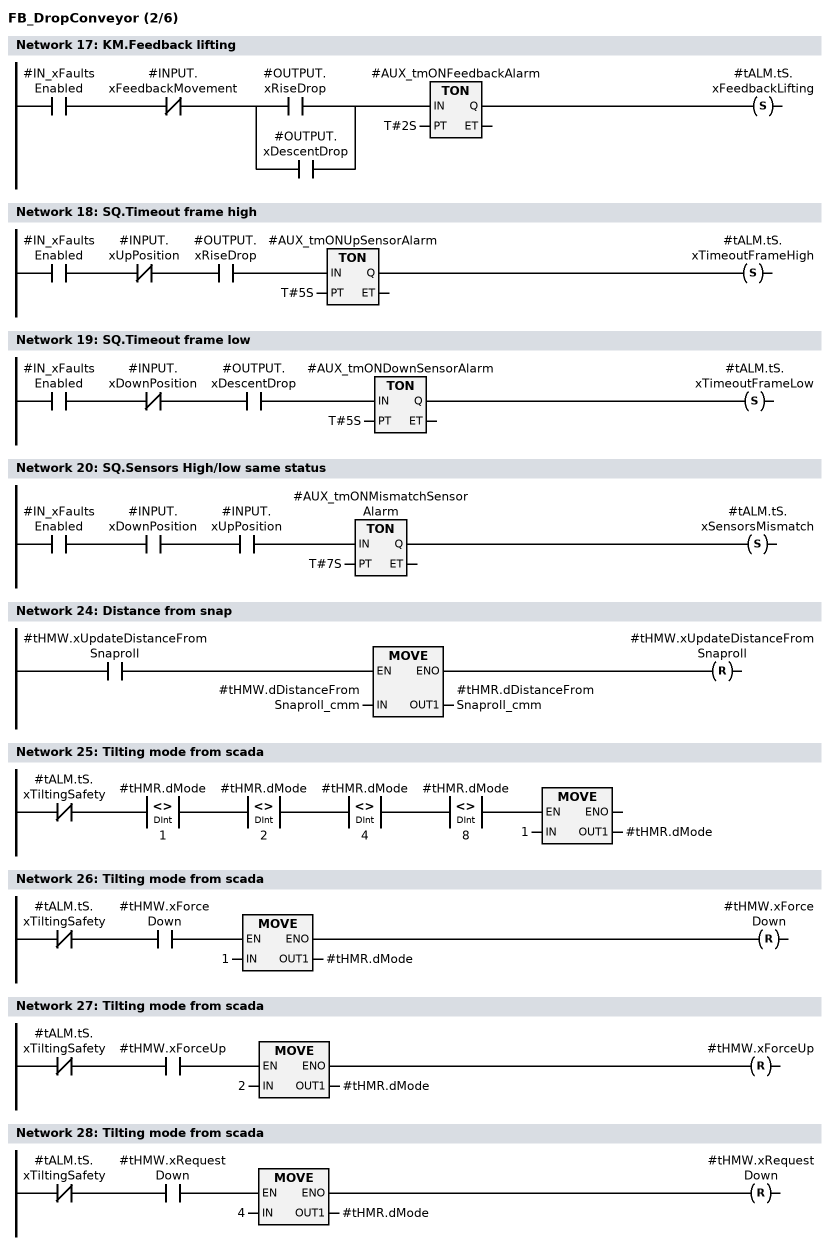
   #AUX_tmONFeedbackAlarm(IN := #IN_xFaultsEnabled AND NOT #INPUT.xFeedbackMovement AND (#OUTPUT.xRiseDrop OR #OUTPUT.xDescentDrop),   // TON
                          PT := T#2S);
   IF #AUX_tmONFeedbackAlarm.Q THEN #tALM.tS.xFeedbackLifting := TRUE; END_IF;
END_REGION

REGION Network 18: SQ.Timeout frame high
   #AUX_tmONUpSensorAlarm(IN := #IN_xFaultsEnabled AND NOT #INPUT.xUpPosition AND #OUTPUT.xRiseDrop, PT := T#5S);   // TON
   IF #AUX_tmONUpSensorAlarm.Q THEN #tALM.tS.xTimeoutFrameHigh := TRUE; END_IF;
END_REGION

REGION Network 19: SQ.Timeout frame low
   #AUX_tmONDownSensorAlarm(IN := #IN_xFaultsEnabled AND NOT #INPUT.xDownPosition AND #OUTPUT.xDescentDrop,   // TON
                           PT := T#5S);
   IF #AUX_tmONDownSensorAlarm.Q THEN #tALM.tS.xTimeoutFrameLow := TRUE; END_IF;
END_REGION

REGION Network 20: SQ.Sensors High/low same status
   #AUX_tmONMismatchSensorAlarm(IN := #IN_xFaultsEnabled AND #INPUT.xDownPosition AND #INPUT.xUpPosition,   // TON
                           PT := T#7S);
   IF #AUX_tmONMismatchSensorAlarm.Q THEN #tALM.tS.xSensorsMismatch := TRUE; END_IF;
END_REGION

REGION Network 21 (SCL): Calculate comulative statuses
       GATHER(IN:=#tALM.tS,
              OUT=>#TMP_dwValue);

       IF #TMP_dwValue <> 0 THEN
           #ST_xStoppingFaults := TRUE;
       ELSE
           #ST_xStoppingFaults := FALSE;
       END_IF;

       GATHER(IN := #tALM.tF,
              OUT => #TMP_dwValue);

       IF #TMP_dwValue <> 0 THEN
           #ST_xFaults := TRUE;
       ELSE
           #ST_xFaults := FALSE;
       END_IF;

       GATHER(IN := #tALM.tW,
              OUT => #TMP_dwValue);

       IF #TMP_dwValue <> 0 THEN
           #ST_xWarnings := TRUE;
       ELSE
           #ST_xWarnings := FALSE;
       END_IF;
END_REGION

REGION Network 22: ### HMI LOGICS ###
END_REGION

REGION Network 23: Break detection
END_REGION

REGION Network 24: Distance from snap
   RUNG wire#powerrail
      Contact( #tHMW.xUpdateDistanceFromSnaproll )
      Move(in := #tHMW.dDistanceFromSnaproll_cmm, out1 => #tHMR.dDistanceFromSnaproll_cmm)
      R_Coil( #tHMW.xUpdateDistanceFromSnaproll )
   END_RUNG
   // the same network as SCL:
   IF #tHMW.xUpdateDistanceFromSnaproll THEN
       #tHMR.dDistanceFromSnaproll_cmm := #tHMW.dDistanceFromSnaproll_cmm;
       #tHMW.xUpdateDistanceFromSnaproll := FALSE;
   END_IF;
END_REGION

REGION Network 25: Tilting mode from scada
   RUNG wire#powerrail
      I_Contact( #tALM.tS.xTiltingSafety )
      { S7_Templates := "SrcType := DInt" } NE_Contact(in1 := #tHMR.dMode, in2 := 1)
      { S7_Templates := "SrcType := DInt" } NE_Contact(in1 := #tHMR.dMode, in2 := 2)
      { S7_Templates := "SrcType := DInt" } NE_Contact(in1 := #tHMR.dMode, in2 := 4)
      { S7_Templates := "SrcType := DInt" } NE_Contact(in1 := #tHMR.dMode, in2 := 8)
      Move(in := 1, out1 => #tHMR.dMode)
   END_RUNG
   // the same network as SCL:
   IF NOT #tALM.tS.xTiltingSafety AND (#tHMR.dMode <> 1) AND (#tHMR.dMode <> 2) AND (#tHMR.dMode <> 4) AND (#tHMR.dMode <> 8) THEN
       #tHMR.dMode := 1;
   END_IF;
END_REGION

REGION Network 26: Tilting mode from scada
   RUNG wire#powerrail
      I_Contact( #tALM.tS.xTiltingSafety )
      Contact( #tHMW.xForceDown )
      Move(in := 1, out1 => #tHMR.dMode)
      R_Coil( #tHMW.xForceDown )
   END_RUNG
   // the same network as SCL:
   IF NOT #tALM.tS.xTiltingSafety AND #tHMW.xForceDown THEN
       #tHMR.dMode := 1;
       #tHMW.xForceDown := FALSE;
   END_IF;
END_REGION

REGION Network 27: Tilting mode from scada
   RUNG wire#powerrail
      I_Contact( #tALM.tS.xTiltingSafety )
      Contact( #tHMW.xForceUp )
      Move(in := 2, out1 => #tHMR.dMode)
      R_Coil( #tHMW.xForceUp )
   END_RUNG
   // the same network as SCL:
   IF NOT #tALM.tS.xTiltingSafety AND #tHMW.xForceUp THEN
       #tHMR.dMode := 2;
       #tHMW.xForceUp := FALSE;
   END_IF;
END_REGION

REGION Network 28: Tilting mode from scada
   RUNG wire#powerrail
      I_Contact( #tALM.tS.xTiltingSafety )
      Contact( #tHMW.xRequestDown )
      Move(in := 4, out1 => #tHMR.dMode)
      R_Coil( #tHMW.xRequestDown )
   END_RUNG
   // the same network as SCL:
   IF NOT #tALM.tS.xTiltingSafety AND #tHMW.xRequestDown THEN
       #tHMR.dMode := 4;
       #tHMW.xRequestDown := FALSE;
   END_IF;
END_REGION

REGION Network 29: Tilting mode from scada
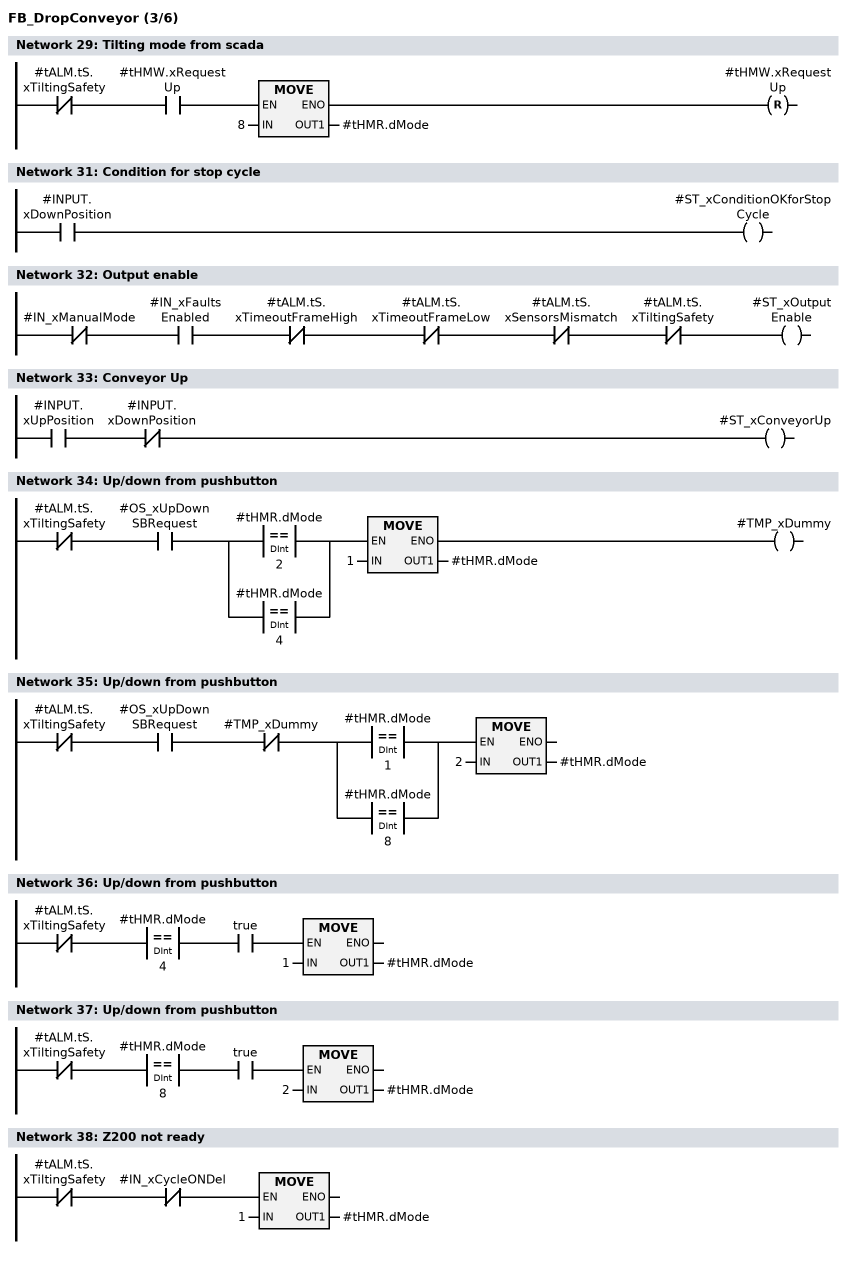
   RUNG wire#powerrail
      I_Contact( #tALM.tS.xTiltingSafety )
      Contact( #tHMW.xRequestUp )
      Move(in := 8, out1 => #tHMR.dMode)
      R_Coil( #tHMW.xRequestUp )
   END_RUNG
   // the same network as SCL:
   IF NOT #tALM.tS.xTiltingSafety AND #tHMW.xRequestUp THEN
       #tHMR.dMode := 8;
       #tHMW.xRequestUp := FALSE;
   END_IF;
END_REGION

REGION Network 30: ### STATUS ###
END_REGION

REGION Network 31: Condition for stop cycle
   RUNG wire#powerrail
      Contact( #INPUT.xDownPosition )
      Coil( #ST_xConditionOKforStopCycle )
   END_RUNG
   // the same network as SCL:
   #ST_xConditionOKforStopCycle := #INPUT.xDownPosition;
END_REGION

REGION Network 32: Output enable
   RUNG wire#powerrail
      I_Contact( #IN_xManualMode )
      Contact( #IN_xFaultsEnabled )
      I_Contact( #tALM.tS.xTimeoutFrameHigh )
      I_Contact( #tALM.tS.xTimeoutFrameLow )
      I_Contact( #tALM.tS.xSensorsMismatch )
      I_Contact( #tALM.tS.xTiltingSafety )
      Coil( #ST_xOutputEnable )
   END_RUNG
   // the same network as SCL:
   #ST_xOutputEnable := NOT #IN_xManualMode AND #IN_xFaultsEnabled AND NOT #tALM.tS.xTimeoutFrameHigh AND NOT #tALM.tS.xTimeoutFrameLow AND NOT #tALM.tS.xSensorsMismatch AND NOT #tALM.tS.xTiltingSafety;
END_REGION

REGION Network 33: Conveyor Up
   RUNG wire#powerrail
      Contact( #INPUT.xUpPosition )
      I_Contact( #INPUT.xDownPosition )
      Coil( #ST_xConveyorUp )
   END_RUNG
   // the same network as SCL:
   #ST_xConveyorUp := #INPUT.xUpPosition AND NOT #INPUT.xDownPosition;
END_REGION

REGION Network 34: Up/down from pushbutton
   RUNG wire#powerrail
      I_Contact( #tALM.tS.xTiltingSafety )
      Contact( #OS_xUpDownSBRequest )
      wire#w1
      { S7_Templates := "SrcType := DInt" } EQ_Contact(in1 := #tHMR.dMode, in2 := 2)
      wire#w2
      Move(in := 1, out1 => #tHMR.dMode)
      Coil( #TMP_xDummy )
   END_RUNG
   RUNG wire#w1
      { S7_Templates := "SrcType := DInt" } EQ_Contact(in1 := #tHMR.dMode, in2 := 4)
   END_RUNG wire#w2
   // the same network as SCL:
   #_w1 := NOT #tALM.tS.xTiltingSafety AND #OS_xUpDownSBRequest AND ((#tHMR.dMode = 2) OR (#tHMR.dMode = 4));
   IF #_w1 THEN #tHMR.dMode := 1; END_IF;
   #TMP_xDummy := #_w1;
END_REGION

REGION Network 35: Up/down from pushbutton
   RUNG wire#powerrail
      I_Contact( #tALM.tS.xTiltingSafety )
      Contact( #OS_xUpDownSBRequest )
      I_Contact( #TMP_xDummy )
      wire#w1
      { S7_Templates := "SrcType := DInt" } EQ_Contact(in1 := #tHMR.dMode, in2 := 1)
      wire#w2
      Move(in := 2, out1 => #tHMR.dMode)
   END_RUNG
   RUNG wire#w1
      { S7_Templates := "SrcType := DInt" } EQ_Contact(in1 := #tHMR.dMode, in2 := 8)
   END_RUNG wire#w2
   // the same network as SCL:
   IF NOT #tALM.tS.xTiltingSafety AND #OS_xUpDownSBRequest AND NOT #TMP_xDummy AND ((#tHMR.dMode = 1) OR (#tHMR.dMode = 8)) THEN
       #tHMR.dMode := 2;
   END_IF;
END_REGION

REGION Network 36: Up/down from pushbutton
   RUNG wire#powerrail
      I_Contact( #tALM.tS.xTiltingSafety )
      { S7_Templates := "SrcType := DInt" } EQ_Contact(in1 := #tHMR.dMode, in2 := 4)
      Contact( true )
      Move(in := 1, out1 => #tHMR.dMode)
   END_RUNG
   // the same network as SCL:
   IF NOT #tALM.tS.xTiltingSafety AND (#tHMR.dMode = 4) AND true THEN #tHMR.dMode := 1; END_IF;
END_REGION

REGION Network 37: Up/down from pushbutton
   RUNG wire#powerrail
      I_Contact( #tALM.tS.xTiltingSafety )
      { S7_Templates := "SrcType := DInt" } EQ_Contact(in1 := #tHMR.dMode, in2 := 8)
      Contact( true )
      Move(in := 2, out1 => #tHMR.dMode)
   END_RUNG
   // the same network as SCL:
   IF NOT #tALM.tS.xTiltingSafety AND (#tHMR.dMode = 8) AND true THEN #tHMR.dMode := 2; END_IF;
END_REGION

REGION Network 38: Z200 not ready
   RUNG wire#powerrail
      I_Contact( #tALM.tS.xTiltingSafety )
      I_Contact( #IN_xCycleONDel )
      Move(in := 1, out1 => #tHMR.dMode)
   END_RUNG
   // the same network as SCL:
   IF NOT #tALM.tS.xTiltingSafety AND NOT #IN_xCycleONDel THEN #tHMR.dMode := 1; END_IF;
END_REGION

REGION Network 39 (SCL): Glass break calculation
   #INO_tRibbon.rgtGlassBreakRequest[#IN_dGlassBreakGetIndex].IN_dDistanceSnaproll_cmm := #tHMR.dDistanceFromSnaproll_cmm;
   #INO_tRibbon.rgtGlassBreakRequest[#IN_dGlassBreakGetIndex].IN_dDownstreamOffset_cmm := #CONST_DBREAKDOWNOFF_CMM;
   #INO_tRibbon.rgtGlassBreakRequest[#IN_dGlassBreakGetIndex].IN_dUpstreamOffset_cmm := #CONST_DBREAKUPOFF_CMM;

   IF #INO_tRibbon.rgtGlassBreakRequest[#IN_dGlassBreakGetIndex].OUT_xDataReady THEN
       #ST_xGlassBreak := #INO_tRibbon.rgtGlassBreakRequest[#IN_dGlassBreakGetIndex].OUT_xGlassBreak;
   END_IF;

   IF #INO_tRibbon.rgtGlassBreakRequest[#IN_dGlassBreakGetIndex].OUT_xDataReady OR NOT #INO_tRibbon.rgtGlassBreakRequest[#IN_dGlassBreakGetIndex].IN_xRequestGlassBreak THEN
       #INO_tRibbon.rgtGlassBreakRequest[#IN_dGlassBreakGetIndex].OUT_xDataReady := FALSE;
       #INO_tRibbon.rgtGlassBreakRequest[#IN_dGlassBreakGetIndex].IN_xRequestGlassBreak := TRUE;
   END_IF;
END_REGION

REGION Network 40: Descent for glass break
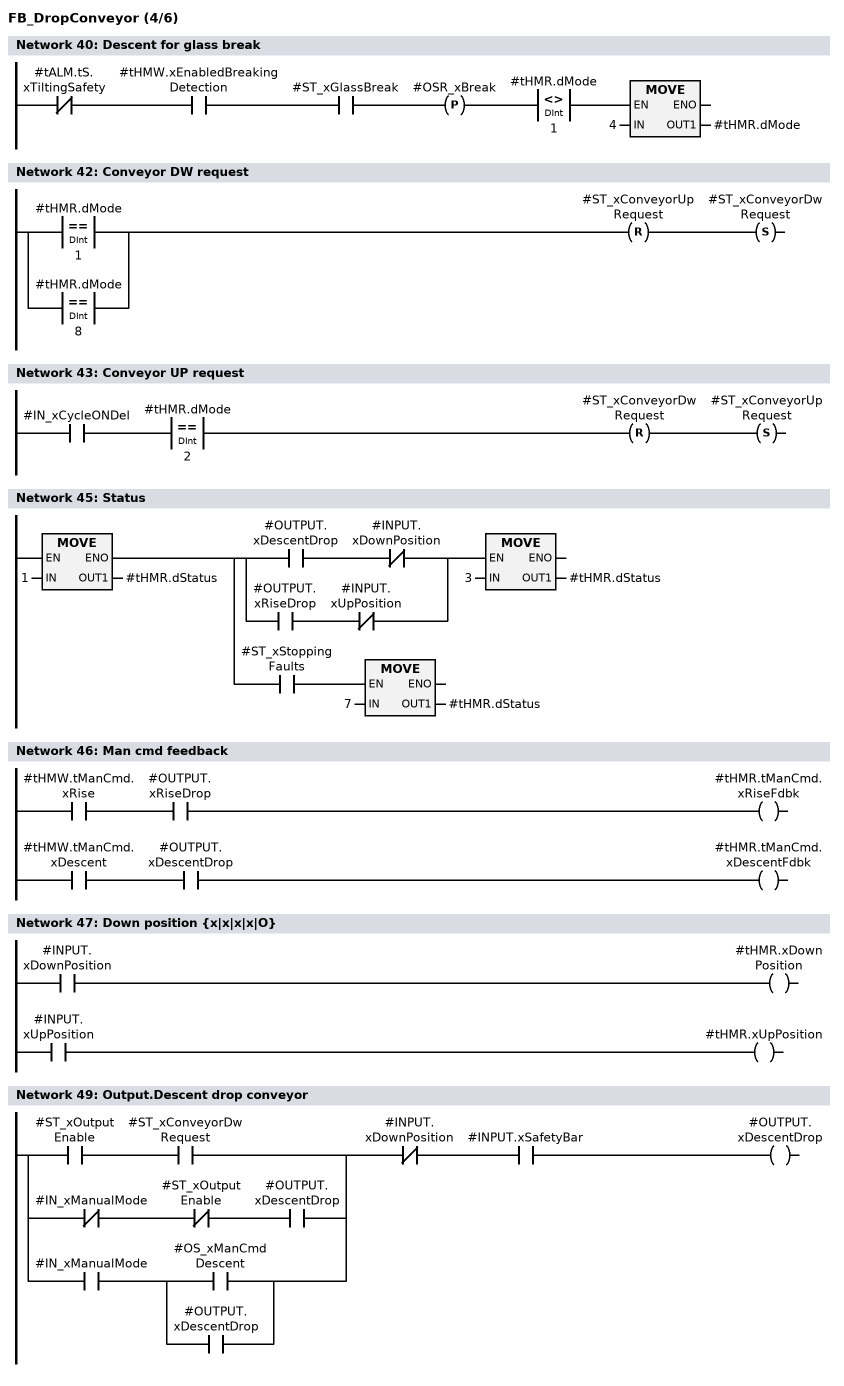
   RUNG wire#powerrail
      I_Contact( #tALM.tS.xTiltingSafety )
      Contact( #tHMW.xEnabledBreakingDetection )
      Contact( #ST_xGlassBreak )
      P_Trig( #OSR_xBreak )
      { S7_Templates := "SrcType := DInt" } NE_Contact(in1 := #tHMR.dMode, in2 := 1)
      Move(in := 4, out1 => #tHMR.dMode)
   END_RUNG
   // the same network as SCL:
   #_w1 := NOT #tALM.tS.xTiltingSafety AND #tHMW.xEnabledBreakingDetection AND #ST_xGlassBreak;
   #_w2 := #_w1 AND NOT #OSR_xBreak;   // rising edge
   #OSR_xBreak := #_w1;
   IF #_w2 AND (#tHMR.dMode <> 1) THEN #tHMR.dMode := 4; END_IF;
END_REGION

REGION Network 41: ### PHASES & LOGICS ###
END_REGION

REGION Network 42: Conveyor DW request
   RUNG wire#powerrail
      { S7_Templates := "SrcType := DInt" } EQ_Contact(in1 := #tHMR.dMode, in2 := 1)
      wire#w1
      R_Coil( #ST_xConveyorUpRequest )
      S_Coil( #ST_xConveyorDwRequest )
   END_RUNG
   RUNG wire#powerrail
      { S7_Templates := "SrcType := DInt" } EQ_Contact(in1 := #tHMR.dMode, in2 := 8)
   END_RUNG wire#w1
   // the same network as SCL:
   IF (#tHMR.dMode = 1) OR (#tHMR.dMode = 8) THEN
       #ST_xConveyorUpRequest := FALSE;
       #ST_xConveyorDwRequest := TRUE;
   END_IF;
END_REGION

REGION Network 43: Conveyor UP request
   RUNG wire#powerrail
      Contact( #IN_xCycleONDel )
      { S7_Templates := "SrcType := DInt" } EQ_Contact(in1 := #tHMR.dMode, in2 := 2)
      R_Coil( #ST_xConveyorDwRequest )
      S_Coil( #ST_xConveyorUpRequest )
   END_RUNG
   // the same network as SCL:
   IF #IN_xCycleONDel AND (#tHMR.dMode = 2) THEN
       #ST_xConveyorDwRequest := FALSE;
       #ST_xConveyorUpRequest := TRUE;
   END_IF;
END_REGION

REGION Network 44: ### HMI STATUS ###
END_REGION

REGION Network 45: Status
   RUNG wire#powerrail
      Move(in := 1, out1 => #tHMR.dStatus)
      wire#w1
      Contact( #OUTPUT.xDescentDrop )
      I_Contact( #INPUT.xDownPosition )
      wire#w2
      Move(in := 3, out1 => #tHMR.dStatus)
   END_RUNG
   RUNG wire#w1
      Contact( #OUTPUT.xRiseDrop )
      I_Contact( #INPUT.xUpPosition )
   END_RUNG wire#w2
   RUNG wire#w1
      Contact( #ST_xStoppingFaults )
      Move(in := 7, out1 => #tHMR.dStatus)
   END_RUNG
   // the same network as SCL:
   #tHMR.dStatus := 1;
   IF (#OUTPUT.xDescentDrop AND NOT #INPUT.xDownPosition) OR (#OUTPUT.xRiseDrop AND NOT #INPUT.xUpPosition) THEN
       #tHMR.dStatus := 3;
   END_IF;
   IF #ST_xStoppingFaults THEN #tHMR.dStatus := 7; END_IF;
END_REGION

REGION Network 46: Man cmd feedback
   RUNG wire#powerrail
      Contact( #tHMW.tManCmd.xRise )
      Contact( #OUTPUT.xRiseDrop )
      Coil( #tHMR.tManCmd.xRiseFdbk )
   END_RUNG
   RUNG wire#powerrail
      Contact( #tHMW.tManCmd.xDescent )
      Contact( #OUTPUT.xDescentDrop )
      Coil( #tHMR.tManCmd.xDescentFdbk )
   END_RUNG
   // the same network as SCL:
   #tHMR.tManCmd.xRiseFdbk := #tHMW.tManCmd.xRise AND #OUTPUT.xRiseDrop;
   #tHMR.tManCmd.xDescentFdbk := #tHMW.tManCmd.xDescent AND #OUTPUT.xDescentDrop;
END_REGION

REGION Network 47: Down position {x|x|x|x|O}
   RUNG wire#powerrail
      Contact( #INPUT.xDownPosition )
      Coil( #tHMR.xDownPosition )
   END_RUNG
   RUNG wire#powerrail
      Contact( #INPUT.xUpPosition )
      Coil( #tHMR.xUpPosition )
   END_RUNG
   // the same network as SCL:
   #tHMR.xDownPosition := #INPUT.xDownPosition;
   #tHMR.xUpPosition := #INPUT.xUpPosition;
END_REGION

REGION Network 48: ### OUTPUT ###
END_REGION

REGION Network 49: Output.Descent drop conveyor
   RUNG wire#powerrail
      Contact( #ST_xOutputEnable )
      Contact( #ST_xConveyorDwRequest )
      wire#w1
      I_Contact( #INPUT.xDownPosition )
      Contact( #INPUT.xSafetyBar )
      Coil( #OUTPUT.xDescentDrop )
   END_RUNG
   RUNG wire#powerrail
      I_Contact( #IN_xManualMode )
      I_Contact( #ST_xOutputEnable )
      Contact( #OUTPUT.xDescentDrop )
   END_RUNG wire#w1
   RUNG wire#powerrail
      Contact( #IN_xManualMode )
      wire#w2
      Contact( #OS_xManCmdDescent )
   END_RUNG wire#w1
   RUNG wire#w2
      Contact( #OUTPUT.xDescentDrop )
   END_RUNG wire#w1
   // the same network as SCL:
   #OUTPUT.xDescentDrop := ((#ST_xOutputEnable AND #ST_xConveyorDwRequest) OR (NOT #IN_xManualMode AND NOT #ST_xOutputEnable AND #OUTPUT.xDescentDrop) OR (#IN_xManualMode AND (#OS_xManCmdDescent OR #OUTPUT.xDescentDrop))) AND NOT #INPUT.xDownPosition AND #INPUT.xSafetyBar;
END_REGION

REGION Network 50: Output.Rise drop conveyor
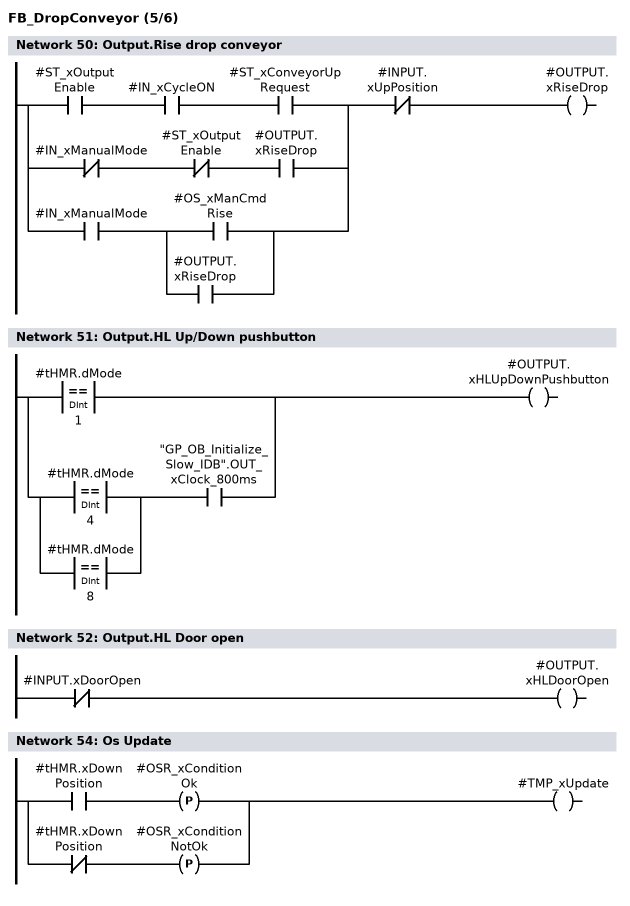
   RUNG wire#powerrail
      Contact( #ST_xOutputEnable )
      Contact( #IN_xCycleON )
      Contact( #ST_xConveyorUpRequest )
      wire#w1
      I_Contact( #INPUT.xUpPosition )
      Coil( #OUTPUT.xRiseDrop )
   END_RUNG
   RUNG wire#powerrail
      I_Contact( #IN_xManualMode )
      I_Contact( #ST_xOutputEnable )
      Contact( #OUTPUT.xRiseDrop )
   END_RUNG wire#w1
   RUNG wire#powerrail
      Contact( #IN_xManualMode )
      wire#w2
      Contact( #OS_xManCmdRise )
   END_RUNG wire#w1
   RUNG wire#w2
      Contact( #OUTPUT.xRiseDrop )
   END_RUNG wire#w1
   // the same network as SCL:
   #OUTPUT.xRiseDrop := ((#ST_xOutputEnable AND #IN_xCycleON AND #ST_xConveyorUpRequest) OR (NOT #IN_xManualMode AND NOT #ST_xOutputEnable AND #OUTPUT.xRiseDrop) OR (#IN_xManualMode AND (#OS_xManCmdRise OR #OUTPUT.xRiseDrop))) AND NOT #INPUT.xUpPosition;
END_REGION

REGION Network 51: Output.HL Up/Down pushbutton
   RUNG wire#powerrail
      { S7_Templates := "SrcType := DInt" } EQ_Contact(in1 := #tHMR.dMode, in2 := 1)
      wire#w1
      Coil( #OUTPUT.xHLUpDownPushbutton )
   END_RUNG
   RUNG wire#powerrail
      { S7_Templates := "SrcType := DInt" } EQ_Contact(in1 := #tHMR.dMode, in2 := 4)
      wire#w2
      Contact( "GP_OB_Initialize_Slow_IDB".OUT_xClock_800ms )
   END_RUNG wire#w1
   RUNG wire#powerrail
      { S7_Templates := "SrcType := DInt" } EQ_Contact(in1 := #tHMR.dMode, in2 := 8)
   END_RUNG wire#w2
   // the same network as SCL:
   #OUTPUT.xHLUpDownPushbutton := (#tHMR.dMode = 1) OR (((#tHMR.dMode = 4) OR (#tHMR.dMode = 8)) AND "GP_OB_Initialize_Slow_IDB".OUT_xClock_800ms);
END_REGION

REGION Network 52: Output.HL Door open
   RUNG wire#powerrail
      I_Contact( #INPUT.xDoorOpen )
      Coil( #OUTPUT.xHLDoorOpen )
   END_RUNG
   // the same network as SCL:
   #OUTPUT.xHLDoorOpen := NOT #INPUT.xDoorOpen;
END_REGION

REGION Network 53: ### REPORT ###
END_REGION

REGION Network 54: Os Update
   RUNG wire#powerrail
      Contact( #tHMR.xDownPosition )
      P_Trig( #OSR_xConditionOk )
      wire#w1
      Coil( #TMP_xUpdate )
   END_RUNG
   RUNG wire#powerrail
      I_Contact( #tHMR.xDownPosition )
      P_Trig( #OSR_xConditionNotOk )
   END_RUNG wire#w1
   // the same network as SCL:
   #_w1 := #tHMR.xDownPosition AND NOT #OSR_xConditionOk;   // rising edge
   #OSR_xConditionOk := #tHMR.xDownPosition;
   #_w2 := NOT #tHMR.xDownPosition AND NOT #OSR_xConditionNotOk;   // rising edge
   #OSR_xConditionNotOk := NOT #tHMR.xDownPosition;
   #TMP_xUpdate := #_w1 OR #_w2;
END_REGION

REGION Network 55: Trap Status
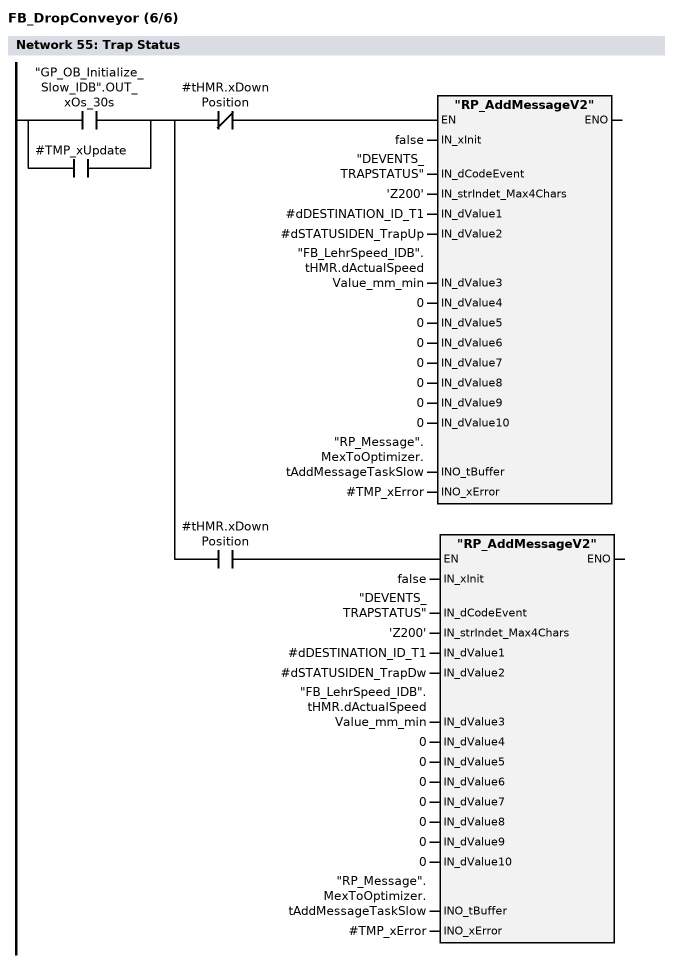
   RUNG wire#powerrail
      Contact( "GP_OB_Initialize_Slow_IDB".OUT_xOs_30s )
      wire#w1
      I_Contact( #tHMR.xDownPosition )
      "RP_AddMessageV2"(IN_xInit := false, IN_dCodeEvent := "DEVENTS_TRAPSTATUS", IN_strIndet_Max4Chars := 'Z200', IN_dValue1 := #dDESTINATION_ID_T1, IN_dValue2 := #dSTATUSIDEN_TrapUp, IN_dValue3 := "FB_LehrSpeed_IDB".tHMR.dActualSpeedValue_mm_min, IN_dValue4 := 0, IN_dValue5 := 0, IN_dValue6 := 0, IN_dValue7 := 0, IN_dValue8 := 0, IN_dValue9 := 0, IN_dValue10 := 0, INO_tBuffer := "RP_Message".MexToOptimizer.tAddMessageTaskSlow, INO_xError := #TMP_xError)
   END_RUNG
   RUNG wire#powerrail
      Contact( #TMP_xUpdate )
   END_RUNG wire#w1
   RUNG wire#w1
      Contact( #tHMR.xDownPosition )
      "RP_AddMessageV2"(IN_xInit := false, IN_dCodeEvent := "DEVENTS_TRAPSTATUS", IN_strIndet_Max4Chars := 'Z200', IN_dValue1 := #dDESTINATION_ID_T1, IN_dValue2 := #dSTATUSIDEN_TrapDw, IN_dValue3 := "FB_LehrSpeed_IDB".tHMR.dActualSpeedValue_mm_min, IN_dValue4 := 0, IN_dValue5 := 0, IN_dValue6 := 0, IN_dValue7 := 0, IN_dValue8 := 0, IN_dValue9 := 0, IN_dValue10 := 0, INO_tBuffer := "RP_Message".MexToOptimizer.tAddMessageTaskSlow, INO_xError := #TMP_xError)
   END_RUNG
   // the same network as SCL:
   #_w1 := "GP_OB_Initialize_Slow_IDB".OUT_xOs_30s OR #TMP_xUpdate;
   IF #_w1 AND NOT #tHMR.xDownPosition THEN
       "RP_AddMessageV2"(IN_xInit := false,
                         IN_dCodeEvent := "DEVENTS_TRAPSTATUS",
                         IN_strIndet_Max4Chars := 'Z200',
                         IN_dValue1 := #dDESTINATION_ID_T1,
                         IN_dValue2 := #dSTATUSIDEN_TrapUp,
                         IN_dValue3 := "FB_LehrSpeed_IDB".tHMR.dActualSpeedValue_mm_min,
                         IN_dValue4 := 0,
                         IN_dValue5 := 0,
                         IN_dValue6 := 0,
                         IN_dValue7 := 0,
                         IN_dValue8 := 0,
                         IN_dValue9 := 0,
                         IN_dValue10 := 0,
                         INO_tBuffer := "RP_Message".MexToOptimizer.tAddMessageTaskSlow,
                         INO_xError := #TMP_xError);
   END_IF;
   IF #_w1 AND #tHMR.xDownPosition THEN
       "RP_AddMessageV2"(IN_xInit := false,
                         IN_dCodeEvent := "DEVENTS_TRAPSTATUS",
                         IN_strIndet_Max4Chars := 'Z200',
                         IN_dValue1 := #dDESTINATION_ID_T1,
                         IN_dValue2 := #dSTATUSIDEN_TrapDw,
                         IN_dValue3 := "FB_LehrSpeed_IDB".tHMR.dActualSpeedValue_mm_min,
                         IN_dValue4 := 0,
                         IN_dValue5 := 0,
                         IN_dValue6 := 0,
                         IN_dValue7 := 0,
                         IN_dValue8 := 0,
                         IN_dValue9 := 0,
                         IN_dValue10 := 0,
                         INO_tBuffer := "RP_Message".MexToOptimizer.tAddMessageTaskSlow,
                         INO_xError := #TMP_xError);
   END_IF;
END_REGION
END_FUNCTION_BLOCK

// folder: 03_Programs_Logics/MCC1201/28_SpeedLehr

FUNCTION_BLOCK "FB_LehrSpeed"   // FB12, LAD
{ S7_Optimized_Access := 'TRUE' }
VERSION : 0.1
   VAR_INPUT
      INPUT_dSpeedSourceEnc1_mm_min : DInt := 0;   // Encoder 1 speed
      INPUT_dSpeedSourceEnc2_mm_min : DInt := 0;   // Encoder 2 speed
      INPUT_dSpeedSourceEth_mm_min : DInt := 0;   // Ethernet speed
      IN_xResetAlarms : Bool;   // Reset alarms
      IN_xEthConnError : Bool;   // Ethernet speed source communication error
   END_VAR
   VAR
      ST_xOutputEnable : Bool := false;   // Output enable
      ST_xPhaseInProgress : Bool := false;   // Phase in progress
      ST_xFaults : Bool := false;   // Cumulative of faults
      ST_xStoppingFaultsEnc1 : Bool := false;   // Cumulative of stopping faults Enc 1
      ST_xStoppingFaultsEnc2 : Bool := false;   // Cumulative of stopping faults Enc 2
      ST_xStoppingFaultsEth : Bool := false;   // Cumulative of stopping faults Eth
      ST_xWarnings : Bool := false;   // Cumulative of warning
      AUX_dLastEthSpeedSourceEnc1_mm_min : DInt := 0;   // Last value of encoder 1 [mm/min]
      AUX_dLastEthSpeedSourceEnc2_mm_min : DInt := 0;   // Last value of encoder 2 [mm/min]
      AUX_dLastEthSpeedSourceEth_mm_min : DInt := 0;   // Last value of ethernet speed [mm/min]
      AUX_dLehrPositionAdvancement : DInt := 0;   // Lehr position advancement [mm/100]
      AUX_tmONTimeoutMessage : TON_TIME;   // Timeout receiving message
   END_VAR
   VAR RETAIN
      tHMR : Struct
         dEncoder1Status : DInt;   // Encoder 1 speed source status (1=Valid 7=Anomaly) {x|x|x|x|O}
         dEncoder1Value_mm_min : DInt;   // Encoder 1 speed source value [mm/min] {mm/min|m/min|x|x|O}
         dEncoder2Status : DInt;   // Encoder 2 speed source status (1=Valid 7=Anomaly) {x|x|x|x|O}
         dEncoder2Value_mm_min : DInt;   // Encoder 2 speed source value [mm/min] {mm/min|m/min|x|x|O}
         dEthStatus : DInt;   // Ethernet speed source status (1=Valid 7=Anomaly) {x|x|x|x|O}
         dEthValue_mm_min : DInt;   // Ethernet speed source value [mm/min] {mm/min|m/min|x|x|O}
         dActualSpeedSource : DInt;   // Actual speed source (1=Manual 2=Encoder_1, 3=Encoder_2, 4=Ethernet)
         dRequestSpeedSource : DInt;   // Request speed source(1=Manual 2=Encoder_1, 3=Encoder_2, 4=Ethernet)
         dActualSpeedValue_mm_min : DInt;   // Actual speed value [mm/min] {mm/min|m/min|x|x|O}
         dActualSpeedValueToConveyor_mm_min : DInt;   // Actual speed value to conveyor [mm/min] {mm/min|m/min|x|x|O}
         dMode : DInt;   // Speed modality (1=Manual;0=Automatic;8=Manual request) {x|x|x|x|O}
      END_STRUCT;
      tHMW : Struct
         dManualSpeedValue_mm_min : DInt;   // Manual speed value [mm/min] {mm/min|m/min|3|22|M}
         xAutoModeReq : Bool;   // Automatic mode request {x|x|x|x|M}
         xManModeReq : Bool;   // Manual mode request {x|x|x|x|M}
         dSpeedOverride_permil : DInt;   // Automatic speed override [‰] {‰|%|-5|5|M}
         dSpeedSelection : DInt;   // Source speed selection (1=Enc1; 2=Enc2; 3=Eth; 4=Auto)
      END_STRUCT;
   END_VAR
   VAR
      tALM : Struct
         tW : Struct   // Warnings
            xSpare_0 : Bool;
            xSpare_1 : Bool;
            xSpare_2 : Bool;
            xSpare_3 : Bool;
            xSpare_4 : Bool;
            xSpare_5 : Bool;
            xSpare_6 : Bool;
            xSpare_7 : Bool;
            xSpare_8 : Bool;
            xSpare_9 : Bool;
            xSpare_10 : Bool;
            xSpare_11 : Bool;
            xSpare_12 : Bool;
            xSpare_13 : Bool;
            xSpare_14 : Bool;
            xSpare_15 : Bool;
            xSpare_16 : Bool;
            xSpare_17 : Bool;
            xSpare_18 : Bool;
            xSpare_19 : Bool;
            xSpare_20 : Bool;
            xSpare_21 : Bool;
            xSpare_22 : Bool;
            xSpare_23 : Bool;
            xSpare_24 : Bool;
            xSpare_25 : Bool;
            xSpare_26 : Bool;
            xSpare_27 : Bool;
            xSpare_28 : Bool;
            xSpare_29 : Bool;
            xSpare_30 : Bool;
            xSpare_31 : Bool;
         END_STRUCT;
         tF : Struct   // Faults
            xSpare_0 : Bool;
            xSpare_1 : Bool;
            xSpare_2 : Bool;
            xSpare_3 : Bool;
            xSpare_4 : Bool;
            xSpare_5 : Bool;
            xSpare_6 : Bool;
            xSpare_7 : Bool;
            xSpare_8 : Bool;
            xSpare_9 : Bool;
            xSpare_10 : Bool;
            xSpare_11 : Bool;
            xSpare_12 : Bool;
            xSpare_13 : Bool;
            xSpare_14 : Bool;
            xSpare_15 : Bool;
            xSpare_16 : Bool;
            xSpare_17 : Bool;
            xSpare_18 : Bool;
            xSpare_19 : Bool;
            xSpare_20 : Bool;
            xSpare_21 : Bool;
            xSpare_22 : Bool;
            xSpare_23 : Bool;
            xSpare_24 : Bool;
            xSpare_25 : Bool;
            xSpare_26 : Bool;
            xSpare_27 : Bool;
            xSpare_28 : Bool;
            xSpare_29 : Bool;
            xSpare_30 : Bool;
            xSpare_31 : Bool;
         END_STRUCT;
         tS : Struct   // Stopping faults
            xEthCommunicationTimeout : Bool;   // Ethernet.Communication timeout
            xEnc1OutOfRange : Bool;   // Ethernet.Enc1 Speed out of range
            xEnc1SpeedDifference : Bool;   // Ethernet.Enc1 Too big speed change
            xEnc2OutOfRange : Bool;   // Ethernet.Enc2 Speed out of range
            xEnc2SpeedDifference : Bool;   // Ethernet.Enc2 Too big speed change
            xEthOutOfRange : Bool;   // Ethernet.Eth Speed out of range
            xEthSpeedDifference : Bool;   // Ethernet.Eth Too big speed change
            xSpare_7 : Bool;
            xSpare_8 : Bool;
            xSpare_9 : Bool;
            xSpare_10 : Bool;
            xSpare_11 : Bool;
            xSpare_12 : Bool;
            xSpare_13 : Bool;
            xSpare_14 : Bool;
            xSpare_15 : Bool;
            xSpare_16 : Bool;
            xSpare_17 : Bool;
            xSpare_18 : Bool;
            xSpare_19 : Bool;
            xSpare_20 : Bool;
            xSpare_21 : Bool;
            xSpare_22 : Bool;
            xSpare_23 : Bool;
            xSpare_24 : Bool;
            xSpare_25 : Bool;
            xSpare_26 : Bool;
            xSpare_27 : Bool;
            xSpare_28 : Bool;
            xSpare_29 : Bool;
            xSpare_30 : Bool;
            xSpare_31 : Bool;
         END_STRUCT;
      END_STRUCT;
   END_VAR
   VAR_TEMP
      TMP_dDummy : DInt;
      TMP_dwValue : DWord;
   END_VAR
   VAR CONSTANT
      CONST_MAX_LEHR_SPEED_MMMIN : DInt := 30000;   // Max lehr speed [mm/min]
      CONST_MIN_LEHR_SPEED_MMMIN : DInt := 100;   // Min lehr speed [mm/min]
   END_VAR
   VAR_TEMP   // added for the SCL form of the ladder/FBD networks
      _w1 : Bool;
   END_VAR
BEGIN

REGION Network 1 (SCL): ### COSTANTS ###
END_REGION

REGION Network 2: ### MATCH ###
END_REGION

REGION Network 3: ####_ALARMS_####
END_REGION

REGION Network 4 (SCL): Reset alarms
   IF #IN_xResetAlarms THEN

       #TMP_dwValue := 0;

       SCATTER(IN:=#TMP_dwValue,
               OUT=>#tALM.tS);

       SCATTER(IN:=#TMP_dwValue,
               OUT=>#tALM.tF);

       SCATTER(IN:=#TMP_dwValue,
               OUT=>#tALM.tW);

   END_IF;
END_REGION

REGION Network 5: Communication error ethernet speed source
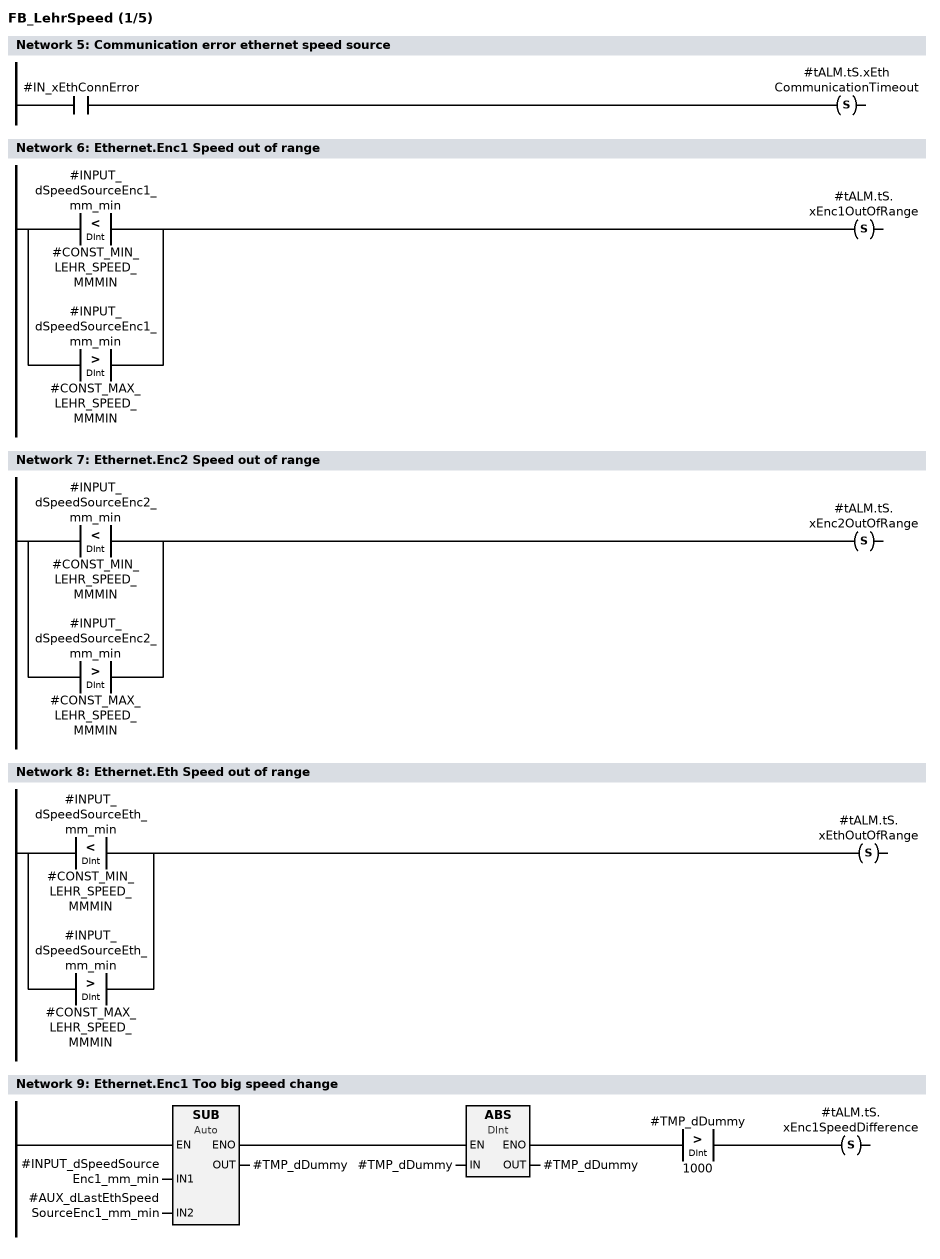
   RUNG wire#powerrail
      Contact( #IN_xEthConnError )
      S_Coil( #tALM.tS.xEthCommunicationTimeout )
   END_RUNG
   // the same network as SCL:
   IF #IN_xEthConnError THEN #tALM.tS.xEthCommunicationTimeout := TRUE; END_IF;
END_REGION

REGION Network 6: Ethernet.Enc1 Speed out of range
   RUNG wire#powerrail
      { S7_Templates := "SrcType := DInt" } LT_Contact(in1 := #INPUT_dSpeedSourceEnc1_mm_min, in2 := #CONST_MIN_LEHR_SPEED_MMMIN)
      wire#w1
      S_Coil( #tALM.tS.xEnc1OutOfRange )
   END_RUNG
   RUNG wire#powerrail
      { S7_Templates := "SrcType := DInt" } GT_Contact(in1 := #INPUT_dSpeedSourceEnc1_mm_min, in2 := #CONST_MAX_LEHR_SPEED_MMMIN)
   END_RUNG wire#w1
   // the same network as SCL:
   IF (#INPUT_dSpeedSourceEnc1_mm_min < #CONST_MIN_LEHR_SPEED_MMMIN) OR (#INPUT_dSpeedSourceEnc1_mm_min > #CONST_MAX_LEHR_SPEED_MMMIN) THEN
       #tALM.tS.xEnc1OutOfRange := TRUE;
   END_IF;
END_REGION

REGION Network 7: Ethernet.Enc2 Speed out of range
   RUNG wire#powerrail
      { S7_Templates := "SrcType := DInt" } LT_Contact(in1 := #INPUT_dSpeedSourceEnc2_mm_min, in2 := #CONST_MIN_LEHR_SPEED_MMMIN)
      wire#w1
      S_Coil( #tALM.tS.xEnc2OutOfRange )
   END_RUNG
   RUNG wire#powerrail
      { S7_Templates := "SrcType := DInt" } GT_Contact(in1 := #INPUT_dSpeedSourceEnc2_mm_min, in2 := #CONST_MAX_LEHR_SPEED_MMMIN)
   END_RUNG wire#w1
   // the same network as SCL:
   IF (#INPUT_dSpeedSourceEnc2_mm_min < #CONST_MIN_LEHR_SPEED_MMMIN) OR (#INPUT_dSpeedSourceEnc2_mm_min > #CONST_MAX_LEHR_SPEED_MMMIN) THEN
       #tALM.tS.xEnc2OutOfRange := TRUE;
   END_IF;
END_REGION

REGION Network 8: Ethernet.Eth Speed out of range
   RUNG wire#powerrail
      { S7_Templates := "SrcType := DInt" } LT_Contact(in1 := #INPUT_dSpeedSourceEth_mm_min, in2 := #CONST_MIN_LEHR_SPEED_MMMIN)
      wire#w1
      S_Coil( #tALM.tS.xEthOutOfRange )
   END_RUNG
   RUNG wire#powerrail
      { S7_Templates := "SrcType := DInt" } GT_Contact(in1 := #INPUT_dSpeedSourceEth_mm_min, in2 := #CONST_MAX_LEHR_SPEED_MMMIN)
   END_RUNG wire#w1
   // the same network as SCL:
   IF (#INPUT_dSpeedSourceEth_mm_min < #CONST_MIN_LEHR_SPEED_MMMIN) OR (#INPUT_dSpeedSourceEth_mm_min > #CONST_MAX_LEHR_SPEED_MMMIN) THEN
       #tALM.tS.xEthOutOfRange := TRUE;
   END_IF;
END_REGION

REGION Network 9: Ethernet.Enc1 Too big speed change
   RUNG wire#powerrail
      Sub(in1 := #INPUT_dSpeedSourceEnc1_mm_min, in2 := #AUX_dLastEthSpeedSourceEnc1_mm_min, out => #TMP_dDummy)
      { S7_Templates := "SrcType := DInt" } Abs(in := #TMP_dDummy, out => #TMP_dDummy)
      { S7_Templates := "SrcType := DInt" } GT_Contact(in1 := #TMP_dDummy, in2 := 1000)
      S_Coil( #tALM.tS.xEnc1SpeedDifference )
   END_RUNG
   // the same network as SCL:
   #TMP_dDummy := #INPUT_dSpeedSourceEnc1_mm_min - #AUX_dLastEthSpeedSourceEnc1_mm_min;
   #TMP_dDummy := ABS(#TMP_dDummy);
   IF #TMP_dDummy > 1000 THEN #tALM.tS.xEnc1SpeedDifference := TRUE; END_IF;
END_REGION

